                 ID := "TC-4011C_MBID",
                 ConnectionType := 11,
                 ActiveEstablished := true,
                 Disconnect := "TC-4011C_W2".Disconnect,
                 MB_Mode := 2,
                 ADDR1 := 192,
                 ADDR2 := 168,
                 ADDR3 := 2,
                 ADDR4 := 20,
                 RemotePort := 502,
                 MB_Unit_ID := 3,
                 MB_Data_Add := 41281,
                 MB_Data_Len := 1,
                 ManualTrigger := NOT "TC-4011C_R1".Processing AND NOT "TC-4011C_R2".Processing AND NOT "TC-4011C_R3".Processing AND NOT "TC-4011C_W1".Processing AND NOT "TC-4011C_W3".Processing AND NOT "TC-4011C_W4".Processing AND NOT "TC-4011C_W2".Processing,
                 MultiFunction := true);
END_REGION

REGION Network 7
   RUNG wire#powerrail
      Contact( "AlwaysFALSE" )
      "AddrMoves"(StartAddr := 41281, EndAddr := 41292, NextAddr := "TC-4011C_W2".Done, Initialize := "TC-4011C_W2".Disconnect, CurrentAddr := "TC-4011A_DB".AddrCtrl.CurrentAddr, Down := "TC-4011A_DB".AddrCtrl.Down, UP := "TC-4011A_DB".AddrCtrl.Up, RisingUp := "TC-4011A_DB".AddrCtrl.RisingUp)
   END_RUNG
   // the same network as SCL:
   IF "AlwaysFALSE" THEN
       "AddrMoves"(StartAddr := 41281,
                   EndAddr := 41292,
                   NextAddr := "TC-4011C_W2".Done,
                   Initialize := "TC-4011C_W2".Disconnect,
                   CurrentAddr := "TC-4011A_DB".AddrCtrl.CurrentAddr,
                   Down := "TC-4011A_DB".AddrCtrl.Down,
                   UP := "TC-4011A_DB".AddrCtrl.Up,
                   RisingUp := "TC-4011A_DB".AddrCtrl.RisingUp);
   END_IF;
END_REGION

REGION Network 8: Write 3
   RUNG wire#powerrail
      "TC-4011C_W3"(ManualTrigger := wire#w1, InterfaceId := 258, ID := "TC-4011C_MBID", ConnectionType := 11, ActiveEstablished := true, Disconnect := "TC-4011C_W3".Disconnect, MB_Mode := 2, ADDR1 := 192, ADDR2 := 168, ADDR3 := 2, ADDR4 := 20, RemotePort := 502, MB_Unit_ID := 3, MB_Data_Add := 41282, MB_Data_Len := 1, MultiFunction := true, Processing =>, Done =>, Busy =>, Error =>, ErrorStatus =>)
   END_RUNG
   RUNG wire#powerrail
      I_Contact( "TC-4011C_R1".Processing )
      I_Contact( "TC-4011C_R2".Processing )
      I_Contact( "TC-4011C_R3".Processing )
      I_Contact( "TC-4011C_W1".Processing )
      I_Contact( "TC-4011C_W2".Processing )
      I_Contact( "TC-4011C_W3".Processing )
      I_Contact( "TC-4011C_W4".Processing )
   END_RUNG wire#w1
   // the same network as SCL:
   "TC-4011C_W3"(InterfaceId := 258,   // "Eurotherm_MB_FB"
                 ID := "TC-4011C_MBID",
                 ConnectionType := 11,
                 ActiveEstablished := true,
                 Disconnect := "TC-4011C_W3".Disconnect,
                 MB_Mode := 2,
                 ADDR1 := 192,
                 ADDR2 := 168,
                 ADDR3 := 2,
                 ADDR4 := 20,
                 RemotePort := 502,
                 MB_Unit_ID := 3,
                 MB_Data_Add := 41282,
                 MB_Data_Len := 1,
                 ManualTrigger := NOT "TC-4011C_R1".Processing AND NOT "TC-4011C_R2".Processing AND NOT "TC-4011C_R3".Processing AND NOT "TC-4011C_W1".Processing AND NOT "TC-4011C_W2".Processing AND NOT "TC-4011C_W3".Processing AND NOT "TC-4011C_W4".Processing,
                 MultiFunction := true);
END_REGION

REGION Network 9: Write 4
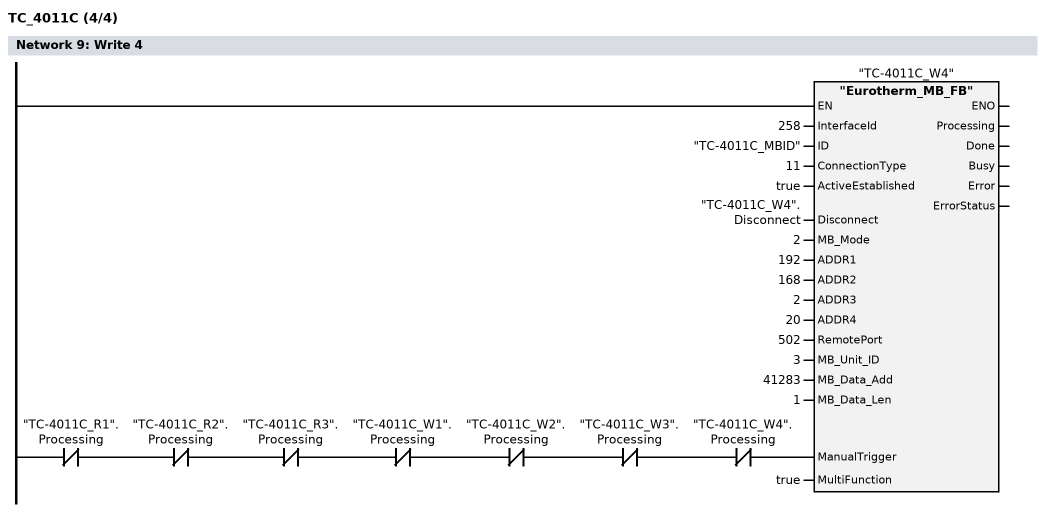
   RUNG wire#powerrail
      "TC-4011C_W4"(ManualTrigger := wire#w1, InterfaceId := 258, ID := "TC-4011C_MBID", ConnectionType := 11, ActiveEstablished := true, Disconnect := "TC-4011C_W4".Disconnect, MB_Mode := 2, ADDR1 := 192, ADDR2 := 168, ADDR3 := 2, ADDR4 := 20, RemotePort := 502, MB_Unit_ID := 3, MB_Data_Add := 41283, MB_Data_Len := 1, MultiFunction := true, Processing =>, Done =>, Busy =>, Error =>, ErrorStatus =>)
   END_RUNG
   RUNG wire#powerrail
      I_Contact( "TC-4011C_R1".Processing )
      I_Contact( "TC-4011C_R2".Processing )
      I_Contact( "TC-4011C_R3".Processing )
      I_Contact( "TC-4011C_W1".Processing )
      I_Contact( "TC-4011C_W2".Processing )
      I_Contact( "TC-4011C_W3".Processing )
      I_Contact( "TC-4011C_W4".Processing )
   END_RUNG wire#w1
   // the same network as SCL:
   "TC-4011C_W4"(InterfaceId := 258,   // "Eurotherm_MB_FB"
                 ID := "TC-4011C_MBID",
                 ConnectionType := 11,
                 ActiveEstablished := true,
                 Disconnect := "TC-4011C_W4".Disconnect,
                 MB_Mode := 2,
                 ADDR1 := 192,
                 ADDR2 := 168,
                 ADDR3 := 2,
                 ADDR4 := 20,
                 RemotePort := 502,
                 MB_Unit_ID := 3,
                 MB_Data_Add := 41283,
                 MB_Data_Len := 1,
                 ManualTrigger := NOT "TC-4011C_R1".Processing AND NOT "TC-4011C_R2".Processing AND NOT "TC-4011C_R3".Processing AND NOT "TC-4011C_W1".Processing AND NOT "TC-4011C_W2".Processing AND NOT "TC-4011C_W3".Processing AND NOT "TC-4011C_W4".Processing,
                 MultiFunction := true);
END_REGION
END_FUNCTION

// folder: Outside Comms/ModBus Comms/Funace_R-402

FUNCTION_BLOCK "YUDIAN_MB_FB"   // FB39, LAD
TITLE = Modbus Block for Real Data Type
{ S7_Optimized_Access := 'TRUE' }
AUTHOR : JL
VERSION : 0.1
   VAR_INPUT
      InterfaceId : Hw_Any;   // HW-identifier of IE-interface submodule
      ID : Conn_Ouc;   // connection reference / identifier
      ConnectionType : Byte;   // type of connection: 11=TCP/IP, 19=UDP (17=TCP/IP)
      ActiveEstablished : Bool := true;   // active/passive connection establishment
      Disconnect : Bool;
      MB_Mode : Byte;
      ADDR1 : Byte;   // IPv4 address
      ADDR2 : Byte;   // IPv4 address
      ADDR3 : Byte;   // IPv4 address
      ADDR4 : Byte;   // IPv4 address
      RemotePort : UInt;   // remote UDP/TCP port number
      MB_Unit_ID : Byte;   // The Modbus slave address
      MB_Data_Add : UDInt;   // Modbus Data Address
      MB_Data_Len : UInt;   // Modbus Data Length
      ManualTrigger : Bool;
      MultiFunction : Bool;   // Depend of the status of the other calls same MB
   END_VAR
   VAR_OUTPUT
      Processing : Bool;
      Done : Bool;
      Busy : Bool;
      Error : Bool;
      ErrorStatus : Word;
   END_VAR
   VAR
      MB_CLIENT_Instance : MB_CLIENT;
      MB_Ctrl : Struct
         REQ : Bool;
         REQ_Again : Bool;
         Disconnect : Bool := false;
         MB_Mode : Byte;   // Modbus Mode
         MB_Data_Address : UDInt;   // Modbus Data Address
         MB_Data_Length : UInt;   // Modbus Data Length
         Connect : TCON_IP_v4;   // Connect Parameters Client
      END_STRUCT;
      MB_Data : Struct
         Buffer : Array[1..16] of Int;
      END_STRUCT;
      "Timer" : Struct
         "1" : IEC_TIMER;
         "2" : IEC_TIMER;
      END_STRUCT;
      OS : Struct
         bit : Array[0..31] of Bool;
      END_STRUCT;
      Process : Struct
         Start : Bool;
         CmdRead : Bool;
         End : Bool;
      END_STRUCT;
   END_VAR
   VAR_TEMP   // added for the SCL form of the ladder/FBD networks
      _w1 : Bool;
      _w2 : Bool;
      _w3 : Bool;
   END_VAR
   // MB_Ctrl.Connect.InterfaceId := 258;
   // MB_Ctrl.Connect.ID := 11;
   // MB_Ctrl.Connect.ConnectionType := 11;
   // MB_Ctrl.Connect.ActiveEstablished := 1;
   // MB_Ctrl.Connect.RemoteAddress.ADDR[1] := 192;
   // MB_Ctrl.Connect.RemoteAddress.ADDR[2] := 168;
   // MB_Ctrl.Connect.RemoteAddress.ADDR[3] := 2;
   // MB_Ctrl.Connect.RemoteAddress.ADDR[4] := 11;
   // MB_Ctrl.Connect.RemotePort := 502;
BEGIN

REGION Network 1 (SCL): Block Parameters
   #MB_Ctrl.Connect.InterfaceId := #InterfaceId;
   #MB_Ctrl.Connect.ID := #ID;
   #MB_Ctrl.Connect.ConnectionType:=#ConnectionType;
   #MB_Ctrl.Disconnect := #Disconnect;
   #MB_Ctrl.MB_Mode:=#MB_Mode;
   #MB_Ctrl.Connect.ActiveEstablished:=#ActiveEstablished;
   #MB_Ctrl.Connect.RemoteAddress.ADDR[1] := #ADDR1;
   #MB_Ctrl.Connect.RemoteAddress.ADDR[2] := #ADDR2;
   #MB_Ctrl.Connect.RemoteAddress.ADDR[3] := #ADDR3;
   #MB_Ctrl.Connect.RemoteAddress.ADDR[4] := #ADDR4;
   #MB_Ctrl.Connect.RemotePort := #RemotePort;
   #MB_CLIENT_Instance.MB_Unit_ID := #MB_Unit_ID;
   #MB_Ctrl.MB_Data_Address := #MB_Data_Add;
   #MB_Ctrl.MB_Data_Length := #MB_Data_Len;
   //#MB_Ctrl.Disconnect := #FbkBusy;
END_REGION

REGION Network 2: Reading Indication
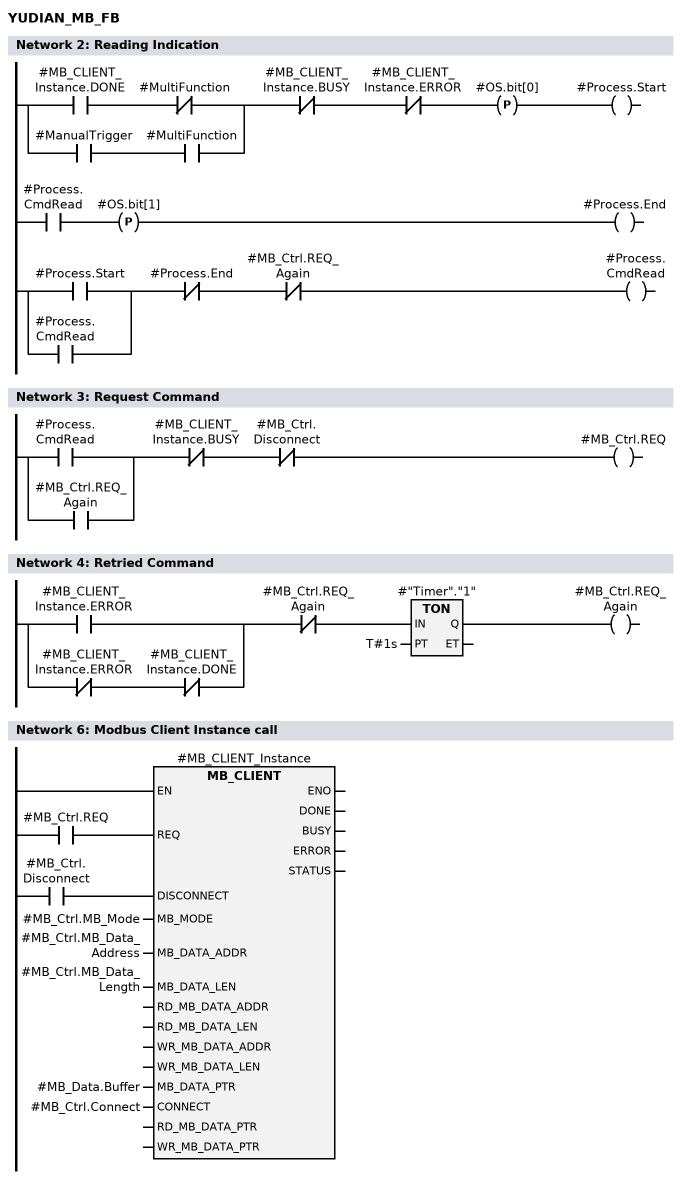
   RUNG wire#powerrail
      Contact( #MB_CLIENT_Instance.DONE )
      I_Contact( #MultiFunction )
      wire#w1
      I_Contact( #MB_CLIENT_Instance.BUSY )
      I_Contact( #MB_CLIENT_Instance.ERROR )
      P_Trig( #OS.bit[0] )
      Coil( #Process.Start )
   END_RUNG
   RUNG wire#powerrail
      Contact( #ManualTrigger )
      Contact( #MultiFunction )
   END_RUNG wire#w1
   RUNG wire#powerrail
      Contact( #Process.CmdRead )
      P_Trig( #OS.bit[1] )
      Coil( #Process.End )
   END_RUNG
   RUNG wire#powerrail
      Contact( #Process.Start )
      wire#w2
      I_Contact( #Process.End )
      I_Contact( #MB_Ctrl.REQ_Again )
      Coil( #Process.CmdRead )
   END_RUNG
   RUNG wire#powerrail
      Contact( #Process.CmdRead )
   END_RUNG wire#w2
   // the same network as SCL:
   #_w1 := ((#MB_CLIENT_Instance.DONE AND NOT #MultiFunction) OR (#ManualTrigger AND #MultiFunction)) AND NOT #MB_CLIENT_Instance.BUSY AND NOT #MB_CLIENT_Instance.ERROR;
   #_w2 := #_w1 AND NOT #OS.bit[0];   // rising edge
   #OS.bit[0] := #_w1;
   #Process.Start := #_w2;
   #_w3 := #Process.CmdRead AND NOT #OS.bit[1];   // rising edge
   #OS.bit[1] := #Process.CmdRead;
   #Process.End := #_w3;
   #Process.CmdRead := (#Process.Start OR #Process.CmdRead) AND NOT #Process.End AND NOT #MB_Ctrl.REQ_Again;
END_REGION

REGION Network 3: Request Command
   RUNG wire#powerrail
      Contact( #Process.CmdRead )
      wire#w1
      I_Contact( #MB_CLIENT_Instance.BUSY )
      I_Contact( #MB_Ctrl.Disconnect )
      Coil( #MB_Ctrl.REQ )
   END_RUNG
   RUNG wire#powerrail
      Contact( #MB_Ctrl.REQ_Again )
   END_RUNG wire#w1
   // the same network as SCL:
   #MB_Ctrl.REQ := (#Process.CmdRead OR #MB_Ctrl.REQ_Again) AND NOT #MB_CLIENT_Instance.BUSY AND NOT #MB_Ctrl.Disconnect;
END_REGION

REGION Network 4: Retried Command
   #"Timer"."1".TON(IN := (#MB_CLIENT_Instance.ERROR OR (NOT #MB_CLIENT_Instance.ERROR AND NOT #MB_CLIENT_Instance.DONE)) AND NOT #MB_Ctrl.REQ_Again,
                    PT := T#1s);
   #MB_Ctrl.REQ_Again := #"Timer"."1".Q;
END_REGION

REGION Network 5 (SCL)
   IF #MB_CLIENT_Instance.ERROR AND #Timer."1".Q THEN
       #MB_CLIENT_Instance.Connected := TRUE;
   END_IF;
END_REGION

REGION Network 6: Modbus Client Instance call
   #MB_CLIENT_Instance(REQ := #MB_Ctrl.REQ,   // MB_CLIENT
                       DISCONNECT := #MB_Ctrl.Disconnect,
                       MB_MODE := #MB_Ctrl.MB_Mode,
                       MB_DATA_ADDR := #MB_Ctrl.MB_Data_Address,
                       MB_DATA_LEN := #MB_Ctrl.MB_Data_Length,
                       MB_DATA_PTR := #MB_Data.Buffer,
                       CONNECT := #MB_Ctrl.Connect);
END_REGION

REGION Network 7 (SCL)
   #Processing := #MB_CLIENT_Instance.BUSY AND NOT #MB_CLIENT_Instance.DONE;
   #Done := #MB_CLIENT_Instance.DONE AND NOT #MB_CLIENT_Instance.BUSY AND NOT #MB_CLIENT_Instance.ERROR;
   #Busy := #MB_CLIENT_Instance.BUSY AND NOT #MB_CLIENT_Instance.DONE;
   #Error := #MB_CLIENT_Instance.ERROR;
   #ErrorStatus := #MB_CLIENT_Instance.STATUS;
END_REGION
END_FUNCTION_BLOCK

// folder: Outside Comms/ModBus Comms/Funace_R-402/TC-402A

FUNCTION "TC_402A" : Void   // FC102, LAD
{ S7_Optimized_Access := 'TRUE' }
VERSION : 0.1
   VAR_TEMP
      MBAddress : UDInt;
      Run : Bool;
      Reset : Bool;
      notProcess : Bool;
   END_VAR
BEGIN

REGION Network 1 (SCL)
   //Data Read 1
   //MOVE_BLK(IN := "Eurothem_Data".Read.Read1.Slaves.Slave1[1],
      //      COUNT := 12,
       //     OUT => "TC-4011A_R1".MB_Data.Buffer[1]);
END_REGION

REGION Network 2
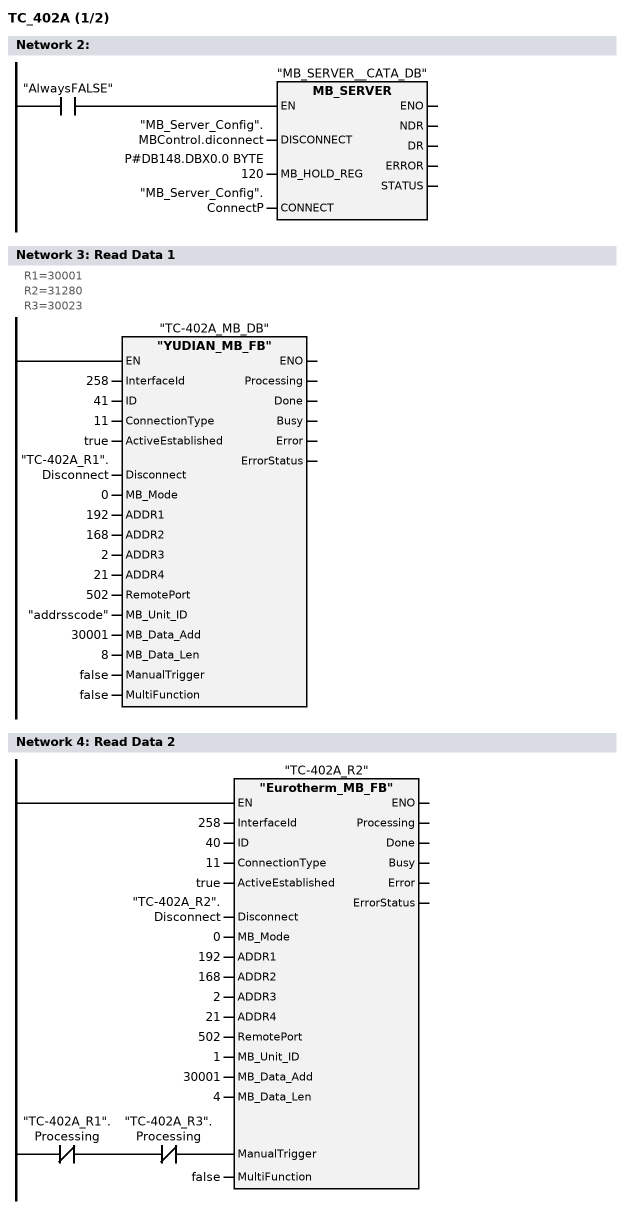
   IF "AlwaysFALSE" THEN
       "MB_SERVER__CATA_DB"(DISCONNECT := "MB_Server_Config".MBControl.diconnect,   // MB_SERVER
                            MB_HOLD_REG := P#DB148.DBX0.0 BYTE 120,
                            CONNECT := "MB_Server_Config".ConnectP);
   END_IF;
END_REGION

REGION Network 3: Read Data 1
   // R1=30001
   // R2=31280
   // R3=30023
   RUNG wire#powerrail
      "TC-402A_MB_DB"(InterfaceId := 258, ID := 41, ConnectionType := 11, ActiveEstablished := true, Disconnect := "TC-402A_R1".Disconnect, MB_Mode := 0, ADDR1 := 192, ADDR2 := 168, ADDR3 := 2, ADDR4 := 21, RemotePort := 502, MB_Unit_ID := "addrsscode", MB_Data_Add := 30001, MB_Data_Len := 8, ManualTrigger := false, MultiFunction := false, Processing =>, Done =>, Busy =>, Error =>, ErrorStatus =>)
   END_RUNG
   // the same network as SCL:
   "TC-402A_MB_DB"(InterfaceId := 258,   // "YUDIAN_MB_FB"
                   ID := 41,
                   ConnectionType := 11,
                   ActiveEstablished := true,
                   Disconnect := "TC-402A_R1".Disconnect,
                   MB_Mode := 0,
                   ADDR1 := 192,
                   ADDR2 := 168,
                   ADDR3 := 2,
                   ADDR4 := 21,
                   RemotePort := 502,
                   MB_Unit_ID := "addrsscode",
                   MB_Data_Add := 30001,
                   MB_Data_Len := 8,
                   ManualTrigger := false,
                   MultiFunction := false);
END_REGION

REGION Network 4: Read Data 2
   RUNG wire#powerrail
      "TC-402A_R2"(ManualTrigger := wire#w1, InterfaceId := 258, ID := 40, ConnectionType := 11, ActiveEstablished := true, Disconnect := "TC-402A_R2".Disconnect, MB_Mode := 0, ADDR1 := 192, ADDR2 := 168, ADDR3 := 2, ADDR4 := 21, RemotePort := 502, MB_Unit_ID := 1, MB_Data_Add := 30001, MB_Data_Len := 4, MultiFunction := false, Processing =>, Done =>, Busy =>, Error =>, ErrorStatus =>)
   END_RUNG
   RUNG wire#powerrail
      I_Contact( "TC-402A_R1".Processing )
      I_Contact( "TC-402A_R3".Processing )
   END_RUNG wire#w1
   // the same network as SCL:
   "TC-402A_R2"(InterfaceId := 258,   // "Eurotherm_MB_FB"
                ID := 40,
                ConnectionType := 11,
                ActiveEstablished := true,
                Disconnect := "TC-402A_R2".Disconnect,
                MB_Mode := 0,
                ADDR1 := 192,
                ADDR2 := 168,
                ADDR3 := 2,
                ADDR4 := 21,
                RemotePort := 502,
                MB_Unit_ID := 1,
                MB_Data_Add := 30001,
                MB_Data_Len := 4,
                ManualTrigger := NOT "TC-402A_R1".Processing AND NOT "TC-402A_R3".Processing,
                MultiFunction := false);
END_REGION

REGION Network 5: Read Data 3
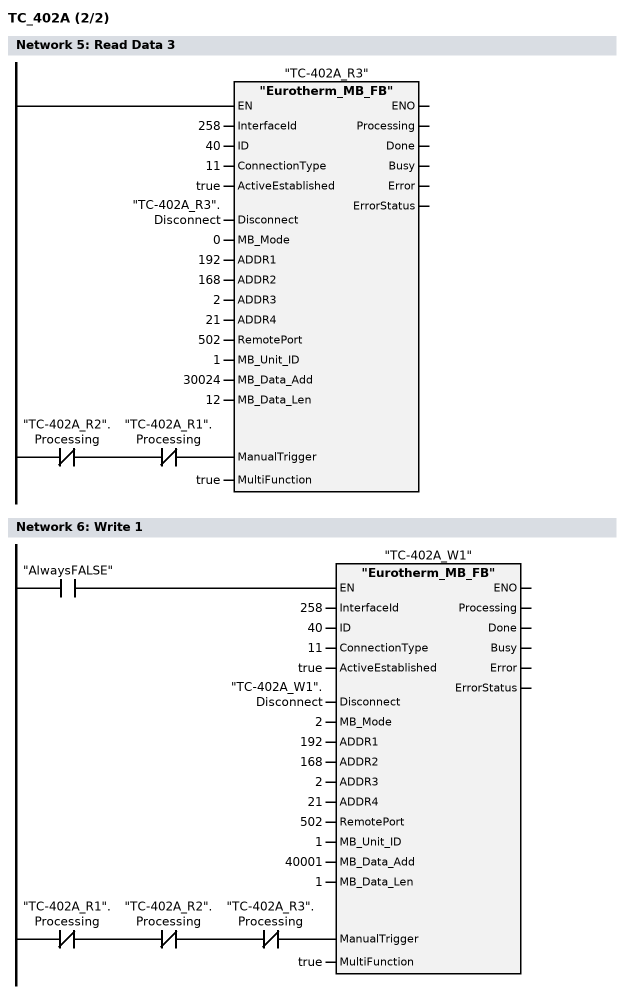
   RUNG wire#powerrail
      "TC-402A_R3"(ManualTrigger := wire#w1, InterfaceId := 258, ID := 40, ConnectionType := 11, ActiveEstablished := true, Disconnect := "TC-402A_R3".Disconnect, MB_Mode := 0, ADDR1 := 192, ADDR2 := 168, ADDR3 := 2, ADDR4 := 21, RemotePort := 502, MB_Unit_ID := 1, MB_Data_Add := 30024, MB_Data_Len := 12, MultiFunction := true, Processing =>, Done =>, Busy =>, Error =>, ErrorStatus =>)
   END_RUNG
   RUNG wire#powerrail
      I_Contact( "TC-402A_R2".Processing )
      I_Contact( "TC-402A_R1".Processing )
   END_RUNG wire#w1
   // the same network as SCL:
   "TC-402A_R3"(InterfaceId := 258,   // "Eurotherm_MB_FB"
                ID := 40,
                ConnectionType := 11,
                ActiveEstablished := true,
                Disconnect := "TC-402A_R3".Disconnect,
                MB_Mode := 0,
                ADDR1 := 192,
                ADDR2 := 168,
                ADDR3 := 2,
                ADDR4 := 21,
                RemotePort := 502,
                MB_Unit_ID := 1,
                MB_Data_Add := 30024,
                MB_Data_Len := 12,
                ManualTrigger := NOT "TC-402A_R2".Processing AND NOT "TC-402A_R1".Processing,
                MultiFunction := true);
END_REGION

REGION Network 6: Write 1
   RUNG wire#powerrail
      Contact( "AlwaysFALSE" )
      "TC-402A_W1"(ManualTrigger := wire#w1, InterfaceId := 258, ID := 40, ConnectionType := 11, ActiveEstablished := true, Disconnect := "TC-402A_W1".Disconnect, MB_Mode := 2, ADDR1 := 192, ADDR2 := 168, ADDR3 := 2, ADDR4 := 21, RemotePort := 502, MB_Unit_ID := 1, MB_Data_Add := 40001, MB_Data_Len := 1, MultiFunction := true, Processing =>, Done =>, Busy =>, Error =>, ErrorStatus =>)
   END_RUNG
   RUNG wire#powerrail
      I_Contact( "TC-402A_R1".Processing )
      I_Contact( "TC-402A_R2".Processing )
      I_Contact( "TC-402A_R3".Processing )
   END_RUNG wire#w1
   // the same network as SCL:
   IF "AlwaysFALSE" THEN
       "TC-402A_W1"(InterfaceId := 258,   // "Eurotherm_MB_FB"
                    ID := 40,
                    ConnectionType := 11,
                    ActiveEstablished := true,
                    Disconnect := "TC-402A_W1".Disconnect,
                    MB_Mode := 2,
                    ADDR1 := 192,
                    ADDR2 := 168,
                    ADDR3 := 2,
                    ADDR4 := 21,
                    RemotePort := 502,
                    MB_Unit_ID := 1,
                    MB_Data_Add := 40001,
                    MB_Data_Len := 1,
                    ManualTrigger := NOT "TC-402A_R1".Processing AND NOT "TC-402A_R2".Processing AND NOT "TC-402A_R3".Processing,
                    MultiFunction := true);
   END_IF;
END_REGION
END_FUNCTION

// folder: Outside Comms/ModBus Comms/Funace_R-402/TC-402B

FUNCTION "TC_402B" : Void   // FC101, LAD
{ S7_Optimized_Access := 'TRUE' }
VERSION : 0.1
   VAR_TEMP
      MBAddress : UDInt;
      Run : Bool;
      Reset : Bool;
      notProcess : Bool;
   END_VAR
BEGIN

REGION Network 1 (SCL)
   //Data Read 1
   //MOVE_BLK(IN := "Eurothem_Data".Read.Read1.Slaves.Slave1[1],
      //      COUNT := 12,
       //     OUT => "TC-4011A_R1".MB_Data.Buffer[1]);
END_REGION

REGION Network 2: Read Data 1
   // R1=30001
   // R2=31280
   // R3=30023
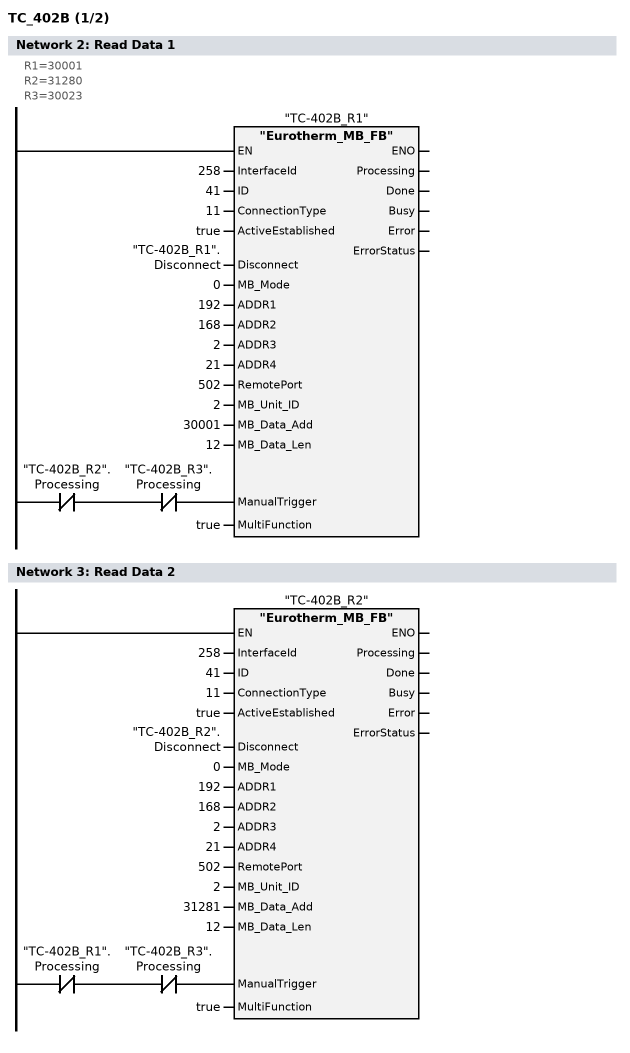
   RUNG wire#powerrail
      "TC-402B_R1"(ManualTrigger := wire#w1, InterfaceId := 258, ID := 41, ConnectionType := 11, ActiveEstablished := true, Disconnect := "TC-402B_R1".Disconnect, MB_Mode := 0, ADDR1 := 192, ADDR2 := 168, ADDR3 := 2, ADDR4 := 21, RemotePort := 502, MB_Unit_ID := 2, MB_Data_Add := 30001, MB_Data_Len := 12, MultiFunction := true, Processing =>, Done =>, Busy =>, Error =>, ErrorStatus =>)
   END_RUNG
   RUNG wire#powerrail
      I_Contact( "TC-402B_R2".Processing )
      I_Contact( "TC-402B_R3".Processing )
   END_RUNG wire#w1
   // the same network as SCL:
   "TC-402B_R1"(InterfaceId := 258,   // "Eurotherm_MB_FB"
                ID := 41,
                ConnectionType := 11,
                ActiveEstablished := true,
                Disconnect := "TC-402B_R1".Disconnect,
                MB_Mode := 0,
                ADDR1 := 192,
                ADDR2 := 168,
                ADDR3 := 2,
                ADDR4 := 21,
                RemotePort := 502,
                MB_Unit_ID := 2,
                MB_Data_Add := 30001,
                MB_Data_Len := 12,
                ManualTrigger := NOT "TC-402B_R2".Processing AND NOT "TC-402B_R3".Processing,
                MultiFunction := true);
END_REGION

REGION Network 3: Read Data 2
   RUNG wire#powerrail
      "TC-402B_R2"(ManualTrigger := wire#w1, InterfaceId := 258, ID := 41, ConnectionType := 11, ActiveEstablished := true, Disconnect := "TC-402B_R2".Disconnect, MB_Mode := 0, ADDR1 := 192, ADDR2 := 168, ADDR3 := 2, ADDR4 := 21, RemotePort := 502, MB_Unit_ID := 2, MB_Data_Add := 31281, MB_Data_Len := 12, MultiFunction := true, Processing =>, Done =>, Busy =>, Error =>, ErrorStatus =>)
   END_RUNG
   RUNG wire#powerrail
      I_Contact( "TC-402B_R1".Processing )
      I_Contact( "TC-402B_R3".Processing )
   END_RUNG wire#w1
   // the same network as SCL:
   "TC-402B_R2"(InterfaceId := 258,   // "Eurotherm_MB_FB"
                ID := 41,
                ConnectionType := 11,
                ActiveEstablished := true,
                Disconnect := "TC-402B_R2".Disconnect,
                MB_Mode := 0,
                ADDR1 := 192,
                ADDR2 := 168,
                ADDR3 := 2,
                ADDR4 := 21,
                RemotePort := 502,
                MB_Unit_ID := 2,
                MB_Data_Add := 31281,
                MB_Data_Len := 12,
                ManualTrigger := NOT "TC-402B_R1".Processing AND NOT "TC-402B_R3".Processing,
                MultiFunction := true);
END_REGION

REGION Network 4: Read Data 3
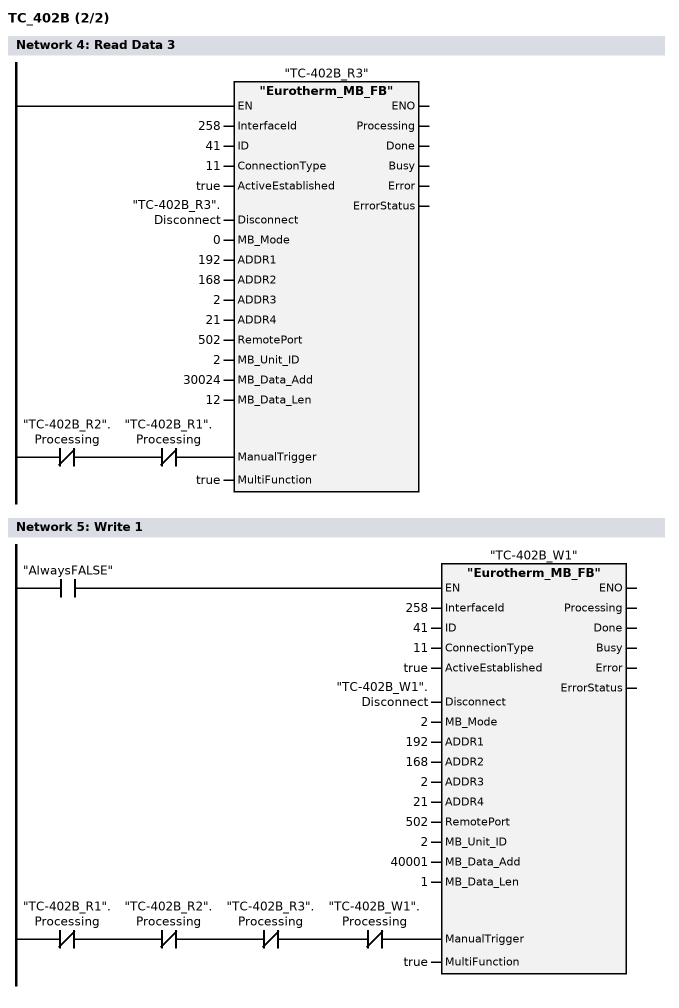
   RUNG wire#powerrail
      "TC-402B_R3"(ManualTrigger := wire#w1, InterfaceId := 258, ID := 41, ConnectionType := 11, ActiveEstablished := true, Disconnect := "TC-402B_R3".Disconnect, MB_Mode := 0, ADDR1 := 192, ADDR2 := 168, ADDR3 := 2, ADDR4 := 21, RemotePort := 502, MB_Unit_ID := 2, MB_Data_Add := 30024, MB_Data_Len := 12, MultiFunction := true, Processing =>, Done =>, Busy =>, Error =>, ErrorStatus =>)
   END_RUNG
   RUNG wire#powerrail
      I_Contact( "TC-402B_R2".Processing )
      I_Contact( "TC-402B_R1".Processing )
   END_RUNG wire#w1
   // the same network as SCL:
   "TC-402B_R3"(InterfaceId := 258,   // "Eurotherm_MB_FB"
                ID := 41,
                ConnectionType := 11,
                ActiveEstablished := true,
                Disconnect := "TC-402B_R3".Disconnect,
                MB_Mode := 0,
                ADDR1 := 192,
                ADDR2 := 168,
                ADDR3 := 2,
                ADDR4 := 21,
                RemotePort := 502,
                MB_Unit_ID := 2,
                MB_Data_Add := 30024,
                MB_Data_Len := 12,
                ManualTrigger := NOT "TC-402B_R2".Processing AND NOT "TC-402B_R1".Processing,
                MultiFunction := true);
END_REGION

REGION Network 5: Write 1
   RUNG wire#powerrail
      Contact( "AlwaysFALSE" )
      "TC-402B_W1"(ManualTrigger := wire#w1, InterfaceId := 258, ID := 41, ConnectionType := 11, ActiveEstablished := true, Disconnect := "TC-402B_W1".Disconnect, MB_Mode := 2, ADDR1 := 192, ADDR2 := 168, ADDR3 := 2, ADDR4 := 21, RemotePort := 502, MB_Unit_ID := 2, MB_Data_Add := 40001, MB_Data_Len := 1, MultiFunction := true, Processing =>, Done =>, Busy =>, Error =>, ErrorStatus =>)
   END_RUNG
   RUNG wire#powerrail
      I_Contact( "TC-402B_R1".Processing )
      I_Contact( "TC-402B_R2".Processing )
      I_Contact( "TC-402B_R3".Processing )
      I_Contact( "TC-402B_W1".Processing )
   END_RUNG wire#w1
   // the same network as SCL:
   IF "AlwaysFALSE" THEN
       "TC-402B_W1"(InterfaceId := 258,   // "Eurotherm_MB_FB"
                    ID := 41,
                    ConnectionType := 11,
                    ActiveEstablished := true,
                    Disconnect := "TC-402B_W1".Disconnect,
                    MB_Mode := 2,
                    ADDR1 := 192,
                    ADDR2 := 168,
                    ADDR3 := 2,
                    ADDR4 := 21,
                    RemotePort := 502,
                    MB_Unit_ID := 2,
                    MB_Data_Add := 40001,
                    MB_Data_Len := 1,
                    ManualTrigger := NOT "TC-402B_R1".Processing AND NOT "TC-402B_R2".Processing AND NOT "TC-402B_R3".Processing AND NOT "TC-402B_W1".Processing,
                    MultiFunction := true);
   END_IF;
END_REGION
END_FUNCTION

// folder: Outside Comms/ModBus Comms/MFCs

FUNCTION_BLOCK "MFC_MB_rDT"   // FB24, LAD
TITLE = Modbus Block for Real Data Type
{ S7_Optimized_Access := 'TRUE' }
AUTHOR : JL
VERSION : 0.1
   VAR_INPUT
      InterfaceId : Hw_Any;   // HW-identifier of IE-interface submodule
      ID : Conn_Ouc;   // connection reference / identifier
      ConnectionType : Byte := 16#11;   // type of connection: 11=TCP/IP, 19=UDP (17=TCP/IP)
      ActiveEstablished : Bool := true;   // active/passive connection establishment
      MB_Mode : Byte;
      ADDR1 : Byte;   // IPv4 address
      ADDR2 : Byte;   // IPv4 address
      ADDR3 : Byte;   // IPv4 address
      ADDR4 : Byte;   // IPv4 address
      RemotePort : UInt := 502;   // remote UDP/TCP port number
      MB_Unit_ID : Byte;   // The Modbus slave address
      MB_Data_Add : UDInt;   // Modbus Data Address in Words (16 bits)
      MB_Data_Len : UInt;   // Modbus Data Length
      FbkBusy : Bool := TRUE;
      MultiFunction : Bool;   // Depend of the status of the other calls same MB
   END_VAR
   VAR_OUTPUT
      Processing : Bool;
      Error : Bool;
   END_VAR
   VAR
      MB_CLIENT_Instance : MB_CLIENT;
      MB_Ctrl : Struct
         REQ : Bool;
         REQ_Again : Bool;
         Disconnect : Bool := false;
         MB_Mode : Byte;   // Modbus Mode
         MB_Data_Address : UDInt;   // Modbus Data Address
         MB_Data_Length : UInt;   // Modbus Data Length
         Connect : TCON_IP_v4;   // Connect Parameters Client
      END_STRUCT;
      MB_Data : Struct
         Buffer : Array[1..8] of Real;
      END_STRUCT;
      "Timer" : Struct
         "1" : IEC_TIMER;
         "2" : IEC_TIMER;
         ConnectionError : IEC_TIMER;
      END_STRUCT;
      OS : Struct
         bit : Array[0..31] of Bool;
      END_STRUCT;
      Process : Struct
         Start : Bool;
         CmdRead : Bool;
         End : Bool;
      END_STRUCT;
   END_VAR
   VAR_TEMP   // added for the SCL form of the ladder/FBD networks
      _w1 : Bool;
      _w2 : Bool;
      _w3 : Bool;
      _w4 : Bool;
   END_VAR
   // MB_Ctrl.Connect.InterfaceId := 258;
   // MB_Ctrl.Connect.ID := 11;
   // MB_Ctrl.Connect.ConnectionType := 11;
   // MB_Ctrl.Connect.ActiveEstablished := 1;
   // MB_Ctrl.Connect.RemoteAddress.ADDR[1] := 192;
   // MB_Ctrl.Connect.RemoteAddress.ADDR[2] := 168;
   // MB_Ctrl.Connect.RemoteAddress.ADDR[3] := 2;
   // MB_Ctrl.Connect.RemoteAddress.ADDR[4] := 11;
   // MB_Ctrl.Connect.RemotePort := 502;
BEGIN

REGION Network 1 (SCL): Block Parameters
   #MB_Ctrl.Connect.InterfaceId := #InterfaceId;
   #MB_Ctrl.Connect.ID := #ID;
   #MB_Ctrl.Connect.ConnectionType:=#ConnectionType;
   #MB_Ctrl.MB_Mode:=#MB_Mode;
   #MB_Ctrl.Connect.ActiveEstablished:=#ActiveEstablished;
   #MB_Ctrl.Connect.RemoteAddress.ADDR[1] := #ADDR1;
   #MB_Ctrl.Connect.RemoteAddress.ADDR[2] := #ADDR2;
   #MB_Ctrl.Connect.RemoteAddress.ADDR[3] := #ADDR3;
   #MB_Ctrl.Connect.RemoteAddress.ADDR[4] := #ADDR4;
   #MB_Ctrl.Connect.RemotePort := #RemotePort;
   #MB_CLIENT_Instance.MB_Unit_ID := #MB_Unit_ID;
   #MB_Ctrl.MB_Data_Address := #MB_Data_Add;
   #MB_Ctrl.MB_Data_Length := #MB_Data_Len;
   //#MB_Ctrl.Disconnect := #FbkBusy;
END_REGION

REGION Network 2: Reading Indication
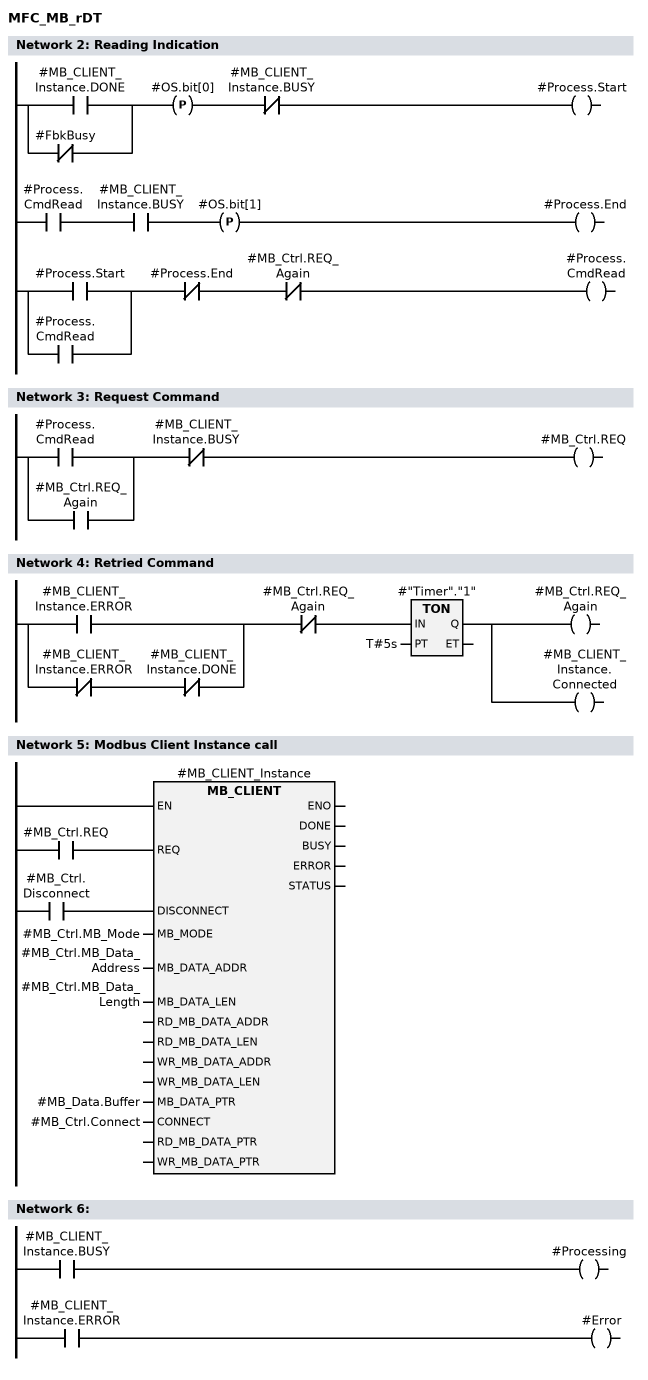
   RUNG wire#powerrail
      Contact( #MB_CLIENT_Instance.DONE )
      wire#w1
      P_Trig( #OS.bit[0] )
      I_Contact( #MB_CLIENT_Instance.BUSY )
      Coil( #Process.Start )
   END_RUNG
   RUNG wire#powerrail
      I_Contact( #FbkBusy )
   END_RUNG wire#w1
   RUNG wire#powerrail
      Contact( #Process.CmdRead )
      Contact( #MB_CLIENT_Instance.BUSY )
      P_Trig( #OS.bit[1] )
      Coil( #Process.End )
   END_RUNG
   RUNG wire#powerrail
      Contact( #Process.Start )
      wire#w2
      I_Contact( #Process.End )
      I_Contact( #MB_Ctrl.REQ_Again )
      Coil( #Process.CmdRead )
   END_RUNG
   RUNG wire#powerrail
      Contact( #Process.CmdRead )
   END_RUNG wire#w2
   // the same network as SCL:
   #_w1 := #MB_CLIENT_Instance.DONE OR NOT #FbkBusy;
   #_w2 := #_w1 AND NOT #OS.bit[0];   // rising edge
   #OS.bit[0] := #_w1;
   #Process.Start := #_w2 AND NOT #MB_CLIENT_Instance.BUSY;
   #_w3 := #Process.CmdRead AND #MB_CLIENT_Instance.BUSY;
   #_w4 := #_w3 AND NOT #OS.bit[1];   // rising edge
   #OS.bit[1] := #_w3;
   #Process.End := #_w4;
   #Process.CmdRead := (#Process.Start OR #Process.CmdRead) AND NOT #Process.End AND NOT #MB_Ctrl.REQ_Again;
END_REGION
